           //"DB323_DM1".DM1[#i].bSt_Tryb.%X12 - Symulacja wejsc urzadzenia: 0-Wylaczona; 1-Zalaczona
           //"DB323_DM1".DM1[#i].bSt_Tryb.%X13 - Praca z wyjsciami urzadzenia: 0-Wylaczona; 1-Zalaczona
           //"DB323_DM1".DM1[#i].bSt_Tryb.%X14 - Stan urzadzenia: 0-Brak odliczania czasu do otwarcia 1-Odliczanie
           //"DB323_DM1".DM1[#i].bSt_Tryb.%X15 - Stan urzadzenia: 0-Brak odliczania czasu do zamkniecia 1-Odliczanie
           //
           //bSt_Urz - STAN - DB323.DBW16 - INT
           //"DB323_DM1".DM1[#i].bSt_Urz.%X0 - STAN(1)- Awaria zbiorcza 1-Aktywna; 0-Brak aktywnosci obiektu
           //"DB323_DM1".DM1[#i].bSt_Urz.%X1 - STAN(2)- Urzadzenie: 1-Zamkniete; 0-Inny stan
           //"DB323_DM1".DM1[#i].bSt_Urz.%X2 - STAN(4)- Urzadzenie: 1-Otwieranie; 0-Inny stan
           //"DB323_DM1".DM1[#i].bSt_Urz.%X3 - STAN(8)- Urzadzenie: 1-Otwarte; 0-Inny stan
           //"DB323_DM1".DM1[#i].bSt_Urz.%X4 - STAN(16)- Urzadzenie: 1-Zamykanie; 0-Inny stan
           //"DB323_DM1".DM1[#i].bSt_Urz.%X5 - STAN(32)- Urzadzenie: 1-Odliczanie czasu zwloki awarii; 0-Inny stan
           //"DB323_DM1".DM1[#i].bSt_Urz.%X6-X7 - STAN- Stan rezerwa
           //
           //bTrP - TRYB PRACY - DB323.DBW17 - INT
           //"DB323_DM1".DM1[#i].bTrP.%X0 - TRYB PRACY(1) - Tryb Remontowy(1): 1-Aktywny; 0-Brak aktywnosci obiektu
           //"DB323_DM1".DM1[#i].bTrP.%X1 - Tryb PRACY(2) - Tryb Sterowania: 1-Lokalny - z szafy; 0-Inny stan
           //"DB323_DM1".DM1[#i].bTrP.%X2 - TRYB PRACY(4) - Tryb Sterowania Zdalnego: 1-Zdalny Reczny; 0-Inny stan
           //"DB323_DM1".DM1[#i].bTrP.%X3 - TRYB PRACY(8) - Tryb Sterowania Zdalnego: 1-Zdalny Automatyczny; 0-Inny stan
           //"DB323_DM1".DM1[#i].bTrP.%X4-X7 - Tryb PRACY(16)(32)(64)(128): Rezerwa
       END_REGION
       REGION Przepisanie danych do obiektu
           "DB323_DM1".DM1[#i].yNrID := #i;
           "DB323_DM1".DM1[#i].yNrPLC := #Nr_Plc;
           "DB323_DM1".DM1[#i].bKier := #bKier;
       END_REGION
       REGION Warunek na wykonanie funkcji
           "DB323_DM1".DM1[#i].bSym.%X0 := "DB323_DM1".DM1[#i].bWeAkt;
           IF "DB323_DM1".DM1[#i].bWeAkt = 0 THEN //Akcja przy deaktywowaniu obiektu
               "DB323_DM1".DM1[#i].bWeAkt := 0;
               "DB323_DM1".DM1[#i].bWeZalAuto := 0;
               "DB323_DM1".DM1[#i].bWePotwZal := 0;
               "DB323_DM1".DM1[#i].bWePotwWyl := 0;
               "DB323_DM1".DM1[#i].bWePotwGot := 0;
               "DB323_DM1".DM1[#i].bWeTrLok := 0;
               "DB323_DM1".DM1[#i].bWeTrRem := 0;
               "DB323_DM1".DM1[#i].bWeAwrZ := 0;
               "DB323_DM1".DM1[#i].bWeBlZmAuto := 0;
               "DB323_DM1".DM1[#i].bWeIlock := 0;
               "DB323_DM1".DM1[#i].bWeKier := 0;
               "DB323_DM1".DM1[#i].bRoZB1 := 0;
               "DB323_DM1".DM1[#i].bRoZB2 := 0;
               "DB323_DM1".DM1[#i].bSym := 0;
               "DB323_DM1".DM1[#i].bSt_Tryb := 0;
               "DB323_DM1".DM1[#i].bSt_Urz := 0;
               "DB323_DM1".DM1[#i].bTrP := 0;
               "DB323_DM1".DM1[#i].bWySter := 0;
               "DB323_DM1".DM1[#i].bWyRst := 0;
               "DB323_DM1".DM1[#i].bWyKier := 0;
           ELSE
               REGION Program funckji
                   REGION Symulacja wejsc - przepisywanie wartosci wejsciowych, gdy nie ma symulacji oprocz bWeAkt
                       IF "DB323_DM1".DM1[#i].bSt_Tryb.%X12 = 0 THEN
                           "DB323_DM1".DM1[#i].bSym.%X1 := "DB323_DM1".DM1[#i].bWeZalAuto;
                           "DB323_DM1".DM1[#i].bSym.%X2 := "DB323_DM1".DM1[#i].bWePotwZal;
                           "DB323_DM1".DM1[#i].bSym.%X3 := "DB323_DM1".DM1[#i].bWePotwWyl;
                           "DB323_DM1".DM1[#i].bSym.%X4 := "DB323_DM1".DM1[#i].bWePotwGot;
                           "DB323_DM1".DM1[#i].bSym.%X5 := "DB323_DM1".DM1[#i].bWeTrLok;
                           "DB323_DM1".DM1[#i].bSym.%X6 := "DB323_DM1".DM1[#i].bWeTrRem;
                           "DB323_DM1".DM1[#i].bSym.%X7 := "DB323_DM1".DM1[#i].bWeAwrZ;
                           "DB323_DM1".DM1[#i].bSym.%X8 := "DB323_DM1".DM1[#i].bWeBlZmAuto;
                           "DB323_DM1".DM1[#i].bSym.%X9 := "DB323_DM1".DM1[#i].bWeIlock;
                           "DB323_DM1".DM1[#i].bSym.%X10 := "DB323_DM1".DM1[#i].bWeKier;
                       END_IF;
                   END_REGION
                   REGION Okreslenie stanow    
                       "DB323_DM1".DM1[#i].bSt_Tryb.%X8 := "DB323_DM1".DM1[#i].bWeAkt;
                       "DB323_DM1".DM1[#i].bSt_Tryb.%X9 := (("DB323_DM1".DM1[#i].bSym.%X8 AND "DB323_DM1".DM1[#i].bSt_Tryb.%X12) OR ("DB323_DM1".DM1[#i].bWeBlZmAuto AND NOT "DB323_DM1".DM1[#i].bSt_Tryb.%X12));
                       "DB323_DM1".DM1[#i].bSt_Tryb.%X11 := (("DB323_DM1".DM1[#i].bSym.%X9 AND "DB323_DM1".DM1[#i].bSt_Tryb.%X12) OR ("DB323_DM1".DM1[#i].bWeIlock AND NOT "DB323_DM1".DM1[#i].bSt_Tryb.%X12));
                       "DB323_DM1".DM1[#i].bSt_Tryb.%X12 := "DB323_DM1".DM1[#i].bRoZB1.%X1;
                       "DB323_DM1".DM1[#i].bSt_Tryb.%X13 := "DB323_DM1".DM1[#i].bRoZB1.%X2;
                       "DB323_DM1".DM1[#i].bSt_Tryb.%X7 := "DB323_DM1".DM1[#i].bRoZB1.%X6;
                   END_REGION
                   REGION Filtracja
                       REGION Timer 1,2 - opoznienie zalaczenia i wylaczenia
                           "DB323_DM1".DM1[#i].bTmr_On_Start := ("DB323_DM1".DM1[#i].bSym.%X1 AND "DB323_DM1".DM1[#i].bSt_Tryb.%X12) OR ("DB323_DM1".DM1[#i].bWeZalAuto AND NOT "DB323_DM1".DM1[#i].bSt_Tryb.%X12) OR ("DB323_DM1".DM1[#i].bRoZB1.%X3 AND NOT "DB323_DM1".DM1[#i].bRoZB1.%X0);
                           "DB323_DM1".DM1[#i].bTmr_Off_Start := NOT "DB323_DM1".DM1[#i].bTmr_On_Start;
                           "FC301_Timer"(iTyp := 1,
                                         bOnOff := "DB323_DM1".DM1[#i].bTmr_On_Start,
                                         bRst := 0,
                                         dCzasZad := "DB323_DM1".DM1[#i].yCzZadOpzZal,
                                         timer_1s := "imp1s",
                                         bOk => "DB323_DM1".DM1[#i].bTmr_On_Ok,
                                         dCzasAkt := "DB323_DM1".DM1[#i].yCzAktOpzZal);
                           "FC301_Timer"(iTyp := 1,
                                         bOnOff := "DB323_DM1".DM1[#i].bTmr_Off_Start,
                                         bRst := 0,
                                         dCzasZad := "DB323_DM1".DM1[#i].yCzZadOpzWyl,
                                         timer_1s := "imp1s",
                                         bOk => "DB323_DM1".DM1[#i].bTmr_Off_Ok,
                                         dCzasAkt := "DB323_DM1".DM1[#i].yCzAktOpzWyl);

                       END_REGION
                       REGION Efekt dzialania timerow 
                           IF "DB323_DM1".DM1[#i].bTmr_On_Ok THEN
                               "DB323_DM1".DM1[#i].bHlp187 := 1;
                           END_IF;
                           IF "DB323_DM1".DM1[#i].bTmr_Off_Ok OR "DB323_DM1".DM1[#i].bSt_Urz = 1 THEN
                               "DB323_DM1".DM1[#i].bHlp187 := 0;
                           END_IF;
                       END_REGION
                       REGION Stany zaworu przy odliczaniu czasu
                           "DB323_DM1".DM1[#i].bSt_Tryb.%X14 := "DB323_DM1".DM1[#i].bTmr_On_Start AND NOT "DB323_DM1".DM1[#i].bTmr_On_Ok;
                           "DB323_DM1".DM1[#i].bSt_Tryb.%X15 := ("DB323_DM1".DM1[#i].bTmr_Off_Start AND NOT "DB323_DM1".DM1[#i].bTmr_Off_Ok);
                       END_REGION
                   END_REGION
                   REGION Generowanie sygnalu alarmu 
                       REGION Zerowanie czasu awarii przy zmianie sterowania podczas ruchu
                           // niepotrzebne a generuje problemy 
                           // "R_TRIG_DB_1"(CLK := "DB323_DM1".DM1[#i].bHlp186 AND "DB323_DM1".DM1[#i].bSt_Urz <> 1,
                           //               Q => "DB323_DM1".DM1[#i].bHlp256);
                           // "R_TRIG_DB_2"(CLK := NOT "DB323_DM1".DM1[#i].bHlp186 AND "DB323_DM1".DM1[#i].bSt_Urz <> 1,
                           //               Q => "DB323_DM1".DM1[#i].bHlp257);
                           // IF "DB323_DM1".DM1[#i].bHlp256 OR "DB323_DM1".DM1[#i].bHlp257 THEN
                           //     "DB323_DM1".DM1[#i].yCzasAktOpzAlm := 0;
                           //    END_IF;
                       END_REGION
                       REGION Sygnal bledu od potwierdzen.
                           // Jezeli brak bitu monitoringu lub bitu pracy z wyjsciami nie ma awarii. Jezeli jest tryb lokalny lub remontowy nie ma awarii

                           "DB323_DM1".DM1[#i].bTmr_Awr_Start := (("DB323_DM1".DM1[#i].bHlp186 XOR (("DB323_DM1".DM1[#i].bWePotwZal AND NOT "DB323_DM1".DM1[#i].bSt_Tryb.%X12) OR ("DB323_DM1".DM1[#i].bSym.%X2 AND "DB323_DM1".DM1[#i].bSt_Tryb.%X12)))
                           OR (NOT "DB323_DM1".DM1[#i].bHlp186 AND NOT (("DB323_DM1".DM1[#i].bWePotwWyl AND NOT "DB323_DM1".DM1[#i].bSt_Tryb.%X12) OR ("DB323_DM1".DM1[#i].bSym.%X3 AND "DB323_DM1".DM1[#i].bSt_Tryb.%X12)))
                           OR ("DB323_DM1".DM1[#i].bHlp186 AND (("DB323_DM1".DM1[#i].bWePotwWyl AND NOT "DB323_DM1".DM1[#i].bSt_Tryb.%X12) OR ("DB323_DM1".DM1[#i].bSym.%X3 AND "DB323_DM1".DM1[#i].bSt_Tryb.%X12)))
                           OR ((("DB323_DM1".DM1[#i].bWePotwZal AND NOT "DB323_DM1".DM1[#i].bSt_Tryb.%X12) OR ("DB323_DM1".DM1[#i].bSym.%X2 AND "DB323_DM1".DM1[#i].bSt_Tryb.%X12))
                           AND (("DB323_DM1".DM1[#i].bWePotwWyl AND NOT "DB323_DM1".DM1[#i].bSt_Tryb.%X12) OR ("DB323_DM1".DM1[#i].bSym.%X3 AND "DB323_DM1".DM1[#i].bSt_Tryb.%X12)))
                           OR (NOT (("DB323_DM1".DM1[#i].bWePotwZal AND NOT "DB323_DM1".DM1[#i].bSt_Tryb.%X12) OR ("DB323_DM1".DM1[#i].bSym.%X2 AND "DB323_DM1".DM1[#i].bSt_Tryb.%X12))
                           AND NOT (("DB323_DM1".DM1[#i].bWePotwWyl AND NOT "DB323_DM1".DM1[#i].bSt_Tryb.%X12) OR ("DB323_DM1".DM1[#i].bSym.%X3 AND "DB323_DM1".DM1[#i].bSt_Tryb.%X12))))
                           AND "DB323_DM1".DM1[#i].bSt_Tryb.%X7 AND "DB323_DM1".DM1[#i].bSt_Tryb.%X13 AND "DB323_DM1".DM1[#i].bTrP <> 1 AND "DB323_DM1".DM1[#i].bTrP <> 2 AND NOT "DB323_DM1".DM1[#i].bRoZB2.%X0;


                       END_REGION
                       REGION Timer 3 - kontrola alarmu
                           "FC301_Timer"(iTyp := 1,
                                         bOnOff := "DB323_DM1".DM1[#i].bTmr_Awr_Start,
                                         bRst := 0,
                                         dCzasZad := "DB323_DM1".DM1[#i].yCzZadOpzAlm,
                                         timer_1s := "imp1s",
                                         bOk => "DB323_DM1".DM1[#i].bTmr_Alm_Ok,
                                         dCzasAkt :="DB323_DM1".DM1[#i].yCzasAktOpzAlm);



                       END_REGION
                       REGION Ustawienie i kasowanie sygnalu awarii
                           IF "DB323_DM1".DM1[#i].bTmr_Alm_Ok THEN
                               "DB323_DM1".DM1[#i].bSt_Tryb.%X0 := 1;
                               "DB323_DM1".DM1[#i].bRoZB1.%X3 := 0;
                               ;
                           END_IF;
                           IF NOT (("DB323_DM1".DM1[#i].bWePotwGot AND NOT "DB323_DM1".DM1[#i].bSt_Tryb.%X12) OR ("DB323_DM1".DM1[#i].bSym.%X4 AND "DB323_DM1".DM1[#i].bSt_Tryb.%X12)) THEN
                               "DB323_DM1".DM1[#i].bSt_Tryb.%X1 := 1
                               ;
                           END_IF;
                           IF ("DB323_DM1".DM1[#i].bWeAwrZ AND NOT "DB323_DM1".DM1[#i].bSt_Tryb.%X12) OR ("DB323_DM1".DM1[#i].bSym.%X7 AND "DB323_DM1".DM1[#i].bSt_Tryb.%X12) THEN
                               "DB323_DM1".DM1[#i].bSt_Tryb.%X2 := 1
                               ;
                           END_IF;
                           IF "DB323_DM1".DM1[#i].bRoZB2.%X0 AND "DB323_DM1".DM1[#i].bSt_Urz = 1 THEN //zmiana 2.10.23 - reset tylko obiektu w awarii
                               "DB323_DM1".DM1[#i].bSt_Tryb := 0
                               ;
                           END_IF;
                       END_REGION
                   END_REGION
                   REGION Tryb pracy i sterowanie wyjsciem
                       REGION Przepisanie potwierdzen na sterowanie reczne gdy tryb lokalny
                           // Przypadek gdy ktos z wlaczonym lokalnie urz. przechodzi na tryb zdalny-reczny
                           IF "DB323_DM1".DM1[#i].bTrP = 2 THEN
                               "DB323_DM1".DM1[#i].bRoZB1.%X0 := 0;

                               IF (("DB323_DM1".DM1[#i].bWePotwWyl AND NOT "DB323_DM1".DM1[#i].bSt_Tryb.%X12) OR ("DB323_DM1".DM1[#i].bSym.%X3 AND "DB323_DM1".DM1[#i].bSt_Tryb.%X12)) THEN
                                   "DB323_DM1".DM1[#i].bRoZB1.%X3 := 0;
                               END_IF;

                               IF (("DB323_DM1".DM1[#i].bWePotwZal AND NOT "DB323_DM1".DM1[#i].bSt_Tryb.%X12) OR ("DB323_DM1".DM1[#i].bSym.%X2 AND "DB323_DM1".DM1[#i].bSt_Tryb.%X12)) THEN
                                   "DB323_DM1".DM1[#i].bRoZB1.%X3 := 1
                                   ;
                               END_IF;
                               ;
                           END_IF;

                       END_REGION
                       REGION Przepisanie potwierdzen na sterowanie reczne gdy tryb zdalny-auto
                           // Przypadek gdy ktos z wlaczonym automatycznie urz. przechodzi na tryb zdalny-reczny
                           IF "DB323_DM1".DM1[#i].bTrP = 8 THEN
                               "DB323_DM1".DM1[#i].bRoZB1.%X3 := (("DB323_DM1".DM1[#i].bWeZalAuto AND NOT "DB323_DM1".DM1[#i].bSt_Tryb.%X12) OR ("DB323_DM1".DM1[#i].bSym.%X1 AND "DB323_DM1".DM1[#i].bSt_Tryb.%X12));
                               "DB323_DM1".DM1[#i].bRoZB1.%X4 := ("DB323_DM1".DM1[#i].bWeKier AND NOT "DB323_DM1".DM1[#i].bSt_Tryb.%X12) OR ("DB323_DM1".DM1[#i].bSym.%X10 AND "DB323_DM1".DM1[#i].bSt_Tryb.%X12);
                           END_IF;

                       END_REGION
                       REGION Blokada zmiany trybu zdalny-automatyczny
                           IF "DB323_DM1".DM1[#i].bTrP = 8 AND "DB323_DM1".DM1[#i].bSt_Tryb.%X9 THEN
                               "DB323_DM1".DM1[#i].bRoZB1.%X0 := 1;
                               ;
                           END_IF;
                       END_REGION
                       REGION Blokada zalaczenia urzadzenia w trybie zdalnym-manualnym przy zalaczonym Interlocku
                           IF "DB323_DM1".DM1[#i].bWeIlock THEN
                               "DB323_DM1".DM1[#i].bRoZB1.%X3 := 0;
                           END_IF;

                       END_REGION

                       REGION Okreslenie trybu pracy wyjscia
                           IF "DB323_DM1".DM1[#i].bRoZB1.%X0 AND NOT "DB323_DM1".DM1[#i].bSt_Tryb.%X9 THEN
                               "DB323_DM1".DM1[#i].bTrP := 8
                               ;
                           END_IF;
                           IF NOT "DB323_DM1".DM1[#i].bRoZB1.%X0 THEN
                               "DB323_DM1".DM1[#i].bTrP := 4
                               ;
                           END_IF;
                           IF ("DB323_DM1".DM1[#i].bWeTrLok AND NOT "DB323_DM1".DM1[#i].bSt_Tryb.%X12) OR ("DB323_DM1".DM1[#i].bSym.%X5 AND "DB323_DM1".DM1[#i].bSt_Tryb.%X12) THEN
                               "DB323_DM1".DM1[#i].bTrP := 2
                               ;
                           END_IF;
                           IF ("DB323_DM1".DM1[#i].bWeTrRem AND NOT "DB323_DM1".DM1[#i].bSt_Tryb.%X12) OR ("DB323_DM1".DM1[#i].bSym.%X6 AND "DB323_DM1".DM1[#i].bSt_Tryb.%X12)THEN
                               "DB323_DM1".DM1[#i].bTrP := 1
                               ;
                           END_IF;
                       END_REGION
                       REGION Sterowanie wyjsciem
                           "DB323_DM1".DM1[#i].bHlp186 := (("DB323_DM1".DM1[#i].bTrP = 8 AND "DB323_DM1".DM1[#i].bHlp187) OR ("DB323_DM1".DM1[#i].bTrP = 4 AND "DB323_DM1".DM1[#i].bRoZB1.%X3 ))
                           AND NOT (("DB323_DM1".DM1[#i].bWeIlock AND NOT "DB323_DM1".DM1[#i].bSt_Tryb.%X12) OR ("DB323_DM1".DM1[#i].bSym.%X9 AND "DB323_DM1".DM1[#i].bSt_Tryb.%X12)) AND "DB323_DM1".DM1[#i].bSt_Urz <> 1;
                           "DB323_DM1".DM1[#i].bWySter := "DB323_DM1".DM1[#i].bHlp186 AND "DB323_DM1". DM1[#i].bSt_Tryb.%X13;
                       END_REGION
                       REGION Sterowanie kierunkiem
                           "DB323_DM1".DM1[#i].bSt_Tryb.%X10 := ("DB323_DM1".DM1[#i].bTrP = 8 AND (("DB323_DM1".DM1[#i].bSym.%X10 AND "DB323_DM1".DM1[#i].bSt_Tryb.%X12) OR ("DB323_DM1".DM1[#i].bWeKier AND NOT "DB323_DM1".DM1[#i].bSt_Tryb.%X12) ))
                           OR ("DB323_DM1".DM1[#i].bTrP = 4 AND "DB323_DM1".DM1[#i].bRoZB1.%X4);
                           "DB323_DM1".DM1[#i].bWyKier := "DB323_DM1".DM1[#i].bSt_Tryb.%X10 AND "DB323_DM1".DM1[#i].bSt_Tryb.%X13;
                       END_REGION
                       REGION Sterowanie resetem
                           "DB323_DM1".DM1[#i].bWyRst := "DB323_DM1".DM1[#i].bRoZB2.%X0;
                       END_REGION
                       REGION Stan urzadzenia
                           //Urzadzenie otwierane
                           //Awaria   
                           IF  "DB323_DM1".DM1[#i].bSt_Tryb.%X0 OR "DB323_DM1".DM1[#i].bSt_Tryb.%X1 OR "DB323_DM1".DM1[#i].bSt_Tryb.%X2 THEN
                               "DB323_DM1".DM1[#i].bSt_Urz := 1;                   

                           //Zamkniete    
                           ELSIF "DB323_DM1".DM1[#i].bTrP <> 2 AND (("DB323_DM1".DM1[#i].bSt_Tryb.%X7 AND "DB323_DM1".DM1[#i].bSt_Tryb.%X13 AND NOT "DB323_DM1".DM1[#i].bHlp186
                               AND (("DB323_DM1".DM1[#i].bWePotwWyl AND NOT "DB323_DM1".DM1[#i].bSt_Tryb.%X12) OR ("DB323_DM1".DM1[#i].bSym.%X3 AND "DB323_DM1".DM1[#i].bSt_Tryb.%X12)) AND NOT ("DB323_DM1".DM1[#i].bWePotwZal OR "DB323_DM1".DM1[#i].bSym.%X2))
                               OR (NOT "DB323_DM1".DM1[#i].bSt_Tryb.%X7 OR NOT "DB323_DM1".DM1[#i].bSt_Tryb.%X13) AND NOT "DB323_DM1".DM1[#i].bHlp186)
                               OR (("DB323_DM1".DM1[#i].bTrP = 2 AND (("DB323_DM1".DM1[#i].bWePotwWyl AND NOT "DB323_DM1".DM1[#i].bSt_Tryb.%X12) OR ("DB323_DM1".DM1[#i].bSym.%X3 AND "DB323_DM1".DM1[#i].bSt_Tryb.%X12))) OR "DB323_DM1".DM1[#i].bTrP = 1) THEN
                               "DB323_DM1".DM1[#i].bSt_Urz := 2;

                           //Otwarte    
                           ELSIF "DB323_DM1".DM1[#i].bTrP <> 2 AND (("DB323_DM1".DM1[#i].bSt_Tryb.%X7 AND "DB323_DM1".DM1[#i].bSt_Tryb.%X13 AND "DB323_DM1".DM1[#i].bHlp186
                               AND NOT (("DB323_DM1".DM1[#i].bWePotwWyl AND NOT "DB323_DM1".DM1[#i].bSt_Tryb.%X12) OR ("DB323_DM1".DM1[#i].bSym.%X3 AND "DB323_DM1".DM1[#i].bSt_Tryb.%X12))
                               AND (("DB323_DM1".DM1[#i].bWePotwZal AND NOT "DB323_DM1".DM1[#i].bSt_Tryb.%X12) OR ("DB323_DM1".DM1[#i].bSym.%X2 AND "DB323_DM1".DM1[#i].bSt_Tryb.%X12)))
                               OR (NOT "DB323_DM1".DM1[#i].bSt_Tryb.%X7 OR NOT "DB323_DM1".DM1[#i].bSt_Tryb.%X13) AND "DB323_DM1".DM1[#i].bHlp186)
                               OR ("DB323_DM1".DM1[#i].bTrP = 2 AND ("DB323_DM1".DM1[#i].bWePotwZal OR "DB323_DM1".DM1[#i].bSym.%X2)) THEN
                               "DB323_DM1".DM1[#i].bSt_Urz := 8;

                           //kazda inna kombinacja potwierdzen niz przy urz. "otwartym"
                           ELSIF "DB323_DM1".DM1[#i].bSt_Tryb.%X7 AND "DB323_DM1".DM1[#i].bSt_Tryb.%X13 AND "DB323_DM1".DM1[#i].bHlp186 THEN
                               "DB323_DM1".DM1[#i].bSt_Urz := 4;

                           //Zamykanie    
                           ELSIF "DB323_DM1".DM1[#i].bSt_Tryb.%X7 AND "DB323_DM1".DM1[#i].bSt_Tryb.%X13 AND NOT "DB323_DM1".DM1[#i].bHlp186 THEN
                               "DB323_DM1".DM1[#i].bSt_Urz := 16;

                           //Brak gotowości    
                           ELSE
                               "DB323_DM1".DM1[#i].bSt_Urz := 0;
                           END_IF;

                       END_REGION
                   END_REGION
                   REGION Ustawienia koncowe
                       // Samokasowanie sygnalow
                       "DB323_DM1".DM1[#i].bRoZB2 := 0;
                       IF "DB323_DM1".DM1[#i].bAoff = 1 THEN
                           "DB323_DM1".DM1[#i].bWeZalAuto := 0;
                           "DB323_DM1".DM1[#i].bWeKier := 0; //27.11.23
                       END_IF;
                   END_REGION
               END_REGION
           END_IF;
       END_REGION
   END_FOR;
END_FUNCTION

FUNCTION "FC331_AI" : Void   // FC331, SCL
{ S7_Optimized_Access := 'TRUE' }
VERSION : 0.1
   VAR_INPUT
      Nr_Ost_Elementu : Int;   // Numer ostatniego elementu, dla ktorego wykonywana jest klasa
      Nr_Plc : Byte;
      Imp_sek : Bool;
   END_VAR
   VAR_TEMP
      i : Int;
   END_VAR
BEGIN
   FOR #i := 1 TO #Nr_Ost_Elementu BY 1 DO
       REGION Opisy bitow sygnalow: bRoz,bSym,bSt,bSt_1,bTrP
           //bRoz - ROZKAZ OPERATORA - DB3331.DBW10 - WORD
           //bRozB1
           //"DB331_AI".AI[#i].bRoZB1.%X0 - Tryb pracy: 0-Zdalny reczny; 1-Zdalny auto
           //"DB331_AI".AI[#i].bRoZB1.%X1 - Symulacja wejsc urz: 0-Wylaczona; 1-Zalaczona
           //"DB331_AI".AI[#i].bRoZB1.%X2 - Rezerwa
           //"DB331_AI".AI[#i].bRoZB1.%X3 - Rezerwa
           //"DB331_AI".AI[#i].bRoZB1.%X4 - Rezerwa
           //"DB331_AI".AI[#i].bRoZB1.%X5 - tryb symulacji pomiaru: 1-zalaczony; 2-wylaczony 
           //"DB331_AI".AI[#i].bRoZB1.%X6-X7 - Rezerwa
           //bRozB2 - impulsy  
           //"DB331_AI".AI[#i].bRoZB2.%X0 - Kasuj awarie (impuls)
           //"DB331_AI".AI[#i].bRoZB2.%X1-X7 - Rezerwa (impuls)
           //
           //bSym - SYM WEJSCIA - DB3331.DBW12 - WORD
           //"DB331_AI".AI[#i].bSym.%X0 - Aktywacja urz. w systemie (u stawiany tylko z programu)
           //"DB331_AI".AI[#i].bSym.%X1 - Rezerwa
           //"DB331_AI".AI[#i].bSym.%X2-X6 - Rezerwa
           //"DB331_AI".AI[#i].bSym.%X7 - Awaria zewnetrzna: 0-Brak; 1-Aktywny
           //"DB331_AI".AI[#i].bSym.%X8 - Blokada zmiany tr. zdalnego z Auto na Man: 0-Brak; 1-Aktywna
           //"DB331_AI".AI[#i].bSym.%X9-X10 - Rezerwa
           //"DB331_AI".AI[#i].bSym.%X11 - W trybie symulacji pomiaru skok w gore o rSymUp / sekunde
           //"DB331_AI".AI[#i].bSym.%X12 - W trybie symulacji pomiaru skok w gore o rSymUp / sekunde
           //"DB331_AI".AI[#i].bSym.%X13-X15 - Rezerwa
           //
           //bSt_Tryb - STAN - DB331.DBW14 - WORD
           //"DB331_AI".AI[#i].bSt_Tryb.%X0 - Awaria toru pomiarowego: 0-Nieaktywna;1-Aktywna
           //"DB331_AI".AI[#i].bSt_Tryb.%X1 - Awaria rezerwa
           //"DB331_AI".AI[#i].bSt_Tryb.%X2 - Awaria zewnetzrna: 0-Nieaktywna; 1-Aktywna
           //"DB331_AI".AI[#i].bSt_Tryb.%X3-X7 - Awaria rezerwa
           //"DB331_AI".AI[#i].bSt_Tryb.%X8 - Urzadzenie aktywowane
           //"DB331_AI".AI[#i].bSt_Tryb.%X9 - Blokada zmaiany tr. zdalnego z Auto na Man: 0-Brak; 1-Aktywna
           //"DB331_AI".AI[#i].bSt_Tryb.%X10-X11 - Awaria rezerwa
           //"DB331_AI".AI[#i].bSt_Tryb.%X12 - Symulacja wejsc urzadzenia: 0-Wylaczona; 1-Zalaczona
           //"DB331_AI".AI[#i].bSt_Tryb.%X13 - Praca z wyjsciami urzadzenia: 0-Wylaczona; 1-Zalaczona
           //"DB331_AI".AI[#i].bSt_Tryb.%X14 - Tryb symulacji pomiaru - z ustawionym sygnalem bWeSymUp lub bWeSymDown
           //"DB331_AI".AI[#i].bSt_Tryb.%X15 - Stan urzadzenia: 0-Brak odliczania czasu do zamkniecia 1-Odliczanie
           //
           //bSt_Urz - STAN - DB331.DBW16 - INT
           //"DB331_AI".AI[#i].bSt_Urz.%X0 - STAN(1)- Awaria zbiorcza 1-Aktywna; 0-Brak aktywnosci obiektu
           //"DB331_AI".AI[#i].bSt_Urz.%X1 - STAN(2)- Przekroczenie gornej granicy alarmowej
           //"DB331_AI".AI[#i].bSt_Urz.%X2 - STAN(4)- Przekroczenie gornej granicy ostrzegawczej
           //"DB331_AI".AI[#i].bSt_Urz.%X3 - STAN(8)- Urzadzenie: 1-Praca normalne; 0-Inny stan
           //"DB331_AI".AI[#i].bSt_Urz.%X4 - STAN(16)- Prog przekroczenia dolnej granicy ostrzegawczej
           //"DB331_AI".AI[#i].bSt_Urz.%X5 - STAN(32)- Prog przekroczenia dolnej granicy alarmowej
           //"DB331_AI".AI[#i].bSt_Urz.%X6-X7 - STAN- Stan rezerwa
           //
           //bTrP - TRYB PRACY - DB331.DBW17 - INT
           //"DB331_AI".AI[#i].bTrP.%X0 - TRYB PRACY(1): 1-Rezerwa; 0-Brak aktywnosci obiektu
           //"DB331_AI".AI[#i].bTrP.%X1 - Tryb PRACY(2): Rezerwa
           //"DB331_AI".AI[#i].bTrP.%X2 - TRYB PRACY(4) - Tryb Sterowania Zdalnego: 1-Zdalny Reczny; 0-Inny stan
           //"DB331_AI".AI[#i].bTrP.%X3 - TRYB PRACY(8) - Tryb Sterowania Zdalnego: 1-Zdalny Automatyczny; 0-Inny stan
           //"DB331_AI".AI[#i].bTrP.%X4-X7 - Tryb PRACY(16)(32)(64)(128): Rezerwa
           //
           //bL - BLOKADA GENEROWANIA ALARMOW - BYTE
           //"DB331_AI".AI[#i].bB.%X0 - PARAMETR - Blokada generowania alarmu HH: 0-Wylaczona; 1-Zalaczona
           //"DB331_AI".AI[#i].bB.%X1 - PARAMETR - Blokada generowania alarmu H: 0-Wylaczona; 1-Zalaczona
           //"DB331_AI".AI[#i].bB.%X2 - PARAMETR - Blokada generowania alarmu L: 0-Wylaczona; 1-Zalaczona
           //"DB331_AI".AI[#i].bB.%X3 - PARAMETR - Blokada generowania alarmu LL: 0-Wylaczona; 1-Zalaczona
           //"DB331_AI".AI[#i].bB.%X4-X7 - Rezerwa
       END_REGION
      REGION Przepisanie danych do obiektu
                  "DB331_AI".AI[#i].yNrID:= #i;
                  "DB331_AI".AI[#i].yNrPLC := #Nr_Plc;
                   END_REGION
      REGION Warunek na wykonanie funkcji
          IF "DB331_AI".AI[#i].bWeAkt = 0 THEN //Akcja przy deaktywowaniu obiektu
                  "DB331_AI".AI[#i].bWeAwrZ := 0;
                  "DB331_AI".AI[#i].bWeBlZmAuto := 0;
                  "DB331_AI".AI[#i].bWeSymUp := 0;
                  "DB331_AI".AI[#i].bWeSymDown := 0;
                  "DB331_AI".AI[#i].bRoZB1 := 0;
                  "DB331_AI".AI[#i].bRoZB2 := 0;
                  "DB331_AI".AI[#i].bSym := 0;
                  "DB331_AI".AI[#i].bSt_Tryb := 0;
                  "DB331_AI".AI[#i].bSt_Urz := 0;
                  "DB331_AI".AI[#i].bTrP := 0;
                  "DB331_AI".AI[#i].bWyRst := 0;

              ELSE
                   REGION Program funkcji
                       REGION Symulacja wejsc - przepisywanie wartosci wejsciowych, gdy nie ma symulacji oprocz bWeAkt
                           IF "DB331_AI".AI[#i].bSt_Tryb.%X12 = 0 THEN
                               "DB331_AI".AI[#i].bSym.%X7 := "DB331_AI".AI[#i].bWeAwrZ;
                               "DB331_AI".AI[#i].bSym.%X8 := "DB331_AI".AI[#i].bWeBlZmAuto;
                               "DB331_AI".AI[#i].bSym.%X11 := "DB331_AI".AI[#i].bWeSymUp;
                               "DB331_AI".AI[#i].bSym.%X12 := "DB331_AI".AI[#i].bWeSymDown;
                           END_IF;
                       END_REGION
                       REGION Okreslenie stanow
                           "DB331_AI".AI[#i].bSt_Tryb.%X8 := "DB331_AI".AI[#i].bWeAkt;
                           "DB331_AI".AI[#i].bSt_Tryb.%X9 := ("DB331_AI".AI[#i].bSym.%X8 AND "DB331_AI".AI[#i].bSt_Tryb.%X12) OR ("DB331_AI".AI[#i].bWeBlZmAuto AND NOT "DB331_AI".AI[#i].bSt_Tryb.%X12);
                           "DB331_AI".AI[#i].bSt_Tryb.%X12 := "DB331_AI".AI[#i].bRoZB1.%X1;
                           "DB331_AI".AI[#i].bSt_Tryb.%X14 := "DB331_AI".AI[#i].bRoZB1.%X5;
                           REGION Blokada zmiany trybu zdalny-automatyczny
                               IF "DB331_AI".AI[#i].bSt_Tryb.%X9 AND "DB331_AI".AI[#i].bTrP.%X3 THEN
                                   "DB331_AI".AI[#i].bRoZB1.%X0 := 1;
                               END_IF;

